screen "信号监控" 800x480, template "按钮"
   TextField "文本域_1" at 237,127 size 39x20; Text '状态'
   TextField "文本域_2" at 348,127 size 39x20; Text '地址'
   TextField "文本域_3" at 573,127 size 73x20; Text '注释名称'
   Group "Group" at 204,122 size 581x341
   TextField "文本域_30" at 240,127 size 39x20; Text '状态'
   Group "Group_1" at 204,122 size 581x341
   SymbolicIOField "符号 I/O 域_1" at 204,71 size 160x35; TextOn '1'; TextOff '0'; TextList "信号监控"
      on Change: ActivateScreenByNumber("跳转画面", 0)
      ProcessValue <- "跳转画面"
   GraphicView "图形视图_2" at 159,127 size 50x50; Picture "图形_2"
   Rectangle "矩形_2" at 207,152 size 109x15
      Appearance <- "操作面板急停"
   Rectangle "矩形_3" at 207,172 size 109x15
      Appearance <- "回原位"
   Rectangle "矩形_4" at 207,193 size 109x15
      Appearance <- "启动按钮"
   Rectangle "矩形_5" at 207,214 size 109x15
      Appearance <- "停止按钮"
   Rectangle "矩形_6" at 207,235 size 109x15
      Appearance <- "手动/自动"
   Rectangle "矩形_7" at 207,256 size 109x15
      Appearance <- "按钮盒急停"
   Rectangle "矩形_8" at 207,277 size 109x15
      Appearance <- "左启动"
   Rectangle "矩形_9" at 207,298 size 109x15
      Appearance <- "右启动"
   Rectangle "矩形_10" at 207,319 size 109x15
      Appearance <- "备用"
   Rectangle "矩形_11" at 207,340 size 109x15
      Appearance <- "安全光幕"
   Rectangle "矩形_12" at 207,361 size 109x15
      Appearance <- "Y1供料器有料"
   Rectangle "矩形_13" at 207,382 size 109x15
      Appearance <- "Y2供料器有料"
   Rectangle "矩形_14" at 207,403 size 109x15
      Appearance <- "1#工装产品信号"
   Rectangle "矩形_15" at 207,424 size 109x15
      Appearance <- "2#工装产品信号"
   TextField "文本域_4" at 348,150 size 41x20; Text 'I0.0'
   TextField "文本域_5" at 348,170 size 41x20; Text 'I0.1'
   TextField "文本域_6" at 348,191 size 41x20; Text 'I0.2'
   TextField "文本域_7" at 348,212 size 41x20; Text 'I0.3'
   TextField "文本域_8" at 348,233 size 41x20; Text 'I0.4'
   TextField "文本域_9" at 348,254 size 41x20; Text 'I0.5'
   TextField "文本域_10" at 348,275 size 41x20; Text 'I0.6'
   TextField "文本域_11" at 348,296 size 41x20; Text 'I0.7'
   TextField "文本域_12" at 348,317 size 41x20; Text 'I1.0'
   TextField "文本域_13" at 348,338 size 41x20; Text 'I1.1'
   TextField "文本域_14" at 348,359 size 41x20; Text 'I1.2'
   TextField "文本域_15" at 348,380 size 41x20; Text 'I1.3'
   TextField "文本域_16" at 348,401 size 41x20; Text 'I1.4'
   TextField "文本域_17" at 348,422 size 41x20; Text 'I1.5'
   TextField "文本域_18" at 561,151 size 101x19; Text '操作面板急停'
   TextField "文本域_19" at 561,171 size 85x19; Text '回原位按钮'
   TextField "文本域_20" at 561,192 size 101x19; Text '面板启动按钮'
   TextField "文本域_21" at 561,213 size 69x19; Text '停止按钮'
   TextField "文本域_22" at 561,234 size 78x19; Text '手动/自动'
   TextField "文本域_23" at 561,255 size 133x19; Text '双手启动面板急停'
   TextField "文本域_24" at 561,276 size 85x19; Text '左启动按钮'
   TextField "文本域_25" at 561,297 size 85x19; Text '右启动按钮'
   TextField "文本域_26" at 561,318 size 37x19; Text '备用'
   TextField "文本域_27" at 561,339 size 69x19; Text '光幕信号'
   TextField "文本域_28" at 561,360 size 103x19; Text 'Y1供料器有料'
   TextField "文本域_29" at 561,381 size 103x19; Text 'Y2供料器有料'
   TextField "文本域_31" at 561,402 size 119x19; Text '工装产品信号1#'
   TextField "文本域_32" at 561,423 size 119x19; Text '工装产品信号2#'

screen "I2.0" 800x480, template "按钮"
   Group "Group_1" at 204,122 size 581x341
   SymbolicIOField "符号 I/O 域_1" at 204,71 size 160x35; TextOn '1'; TextOff '0'; TextList "信号监控"
      on Change: ActivateScreenByNumber("跳转画面", 0)
      ProcessValue <- "跳转画面"
   GraphicView "图形视图_2" at 159,127 size 50x50; Picture "图形_2"
   Rectangle "矩形_2" at 207,152 size 109x15
      Appearance <- "气夹气缸到位2"
   Rectangle "矩形_3" at 207,172 size 109x15
      Appearance <- "气夹气缸到位1"
   Rectangle "矩形_4" at 207,193 size 109x15
      Appearance <- "工具错误"
   Rectangle "矩形_5" at 207,214 size 109x15
      Appearance <- "工具拧紧OK"
   Rectangle "矩形_6" at 207,235 size 109x15
      Appearance <- "工具拧紧NG"
   Rectangle "矩形_7" at 207,256 size 109x15
      Appearance <- "工具准备好"
   Rectangle "矩形_8" at 207,277 size 109x15
      Appearance <- "工具运行"
   Rectangle "矩形_9" at 207,298 size 109x15
      Appearance <- "气源压力检测"
   TextField "文本域_4" at 348,150 size 41x20; Text 'I2.0'
   TextField "文本域_5" at 348,170 size 41x20; Text 'I2.1'
   TextField "文本域_6" at 348,191 size 41x20; Text 'I2.2'
   TextField "文本域_7" at 348,212 size 41x20; Text 'I2.3'
   TextField "文本域_8" at 348,233 size 41x20; Text 'I2.4'
   TextField "文本域_9" at 348,254 size 41x20; Text 'I2.5'
   TextField "文本域_10" at 348,275 size 41x20; Text 'I2.6'
   TextField "文本域_11" at 348,296 size 41x20; Text 'I2.7'
   TextField "文本域_18" at 561,151 size 110x19; Text '气缸气夹到位2'
   TextField "文本域_19" at 561,171 size 110x19; Text '气缸气夹到位1'
   TextField "文本域_20" at 561,192 size 69x19; Text '工具错误'
   TextField "文本域_21" at 561,213 size 87x19; Text '工具拧紧OK'
   TextField "文本域_22" at 561,234 size 87x19; Text '工具拧紧NG'
   TextField "文本域_23" at 561,255 size 85x19; Text '工具准备好'
   TextField "文本域_24" at 561,276 size 69x19; Text '工具运行'
   TextField "文本域_25" at 561,297 size 101x19; Text '气源压力检测'
   Group "Group" at 204,122 size 581x341
   TextField "文本域_30" at 240,127 size 39x20; Text '状态'
   TextField "文本域_1" at 237,127 size 39x20; Text '状态'
   TextField "文本域_2" at 348,127 size 39x20; Text '地址'
   TextField "文本域_3" at 573,127 size 73x20; Text '注释名称'

screen "I3.0" 800x480, template "按钮"
   Group "Group_1" at 204,122 size 581x341
   SymbolicIOField "符号 I/O 域_1" at 204,71 size 160x35; TextOn '1'; TextOff '0'; TextList "信号监控"
      on Change: ActivateScreenByNumber("跳转画面", 0)
      ProcessValue <- "跳转画面"
   GraphicView "图形视图_2" at 159,127 size 50x50; Picture "图形_2"
   Rectangle "矩形_2" at 207,152 size 109x15
      Appearance <- "光栅屏蔽对射开关"
   Rectangle "矩形_3" at 207,172 size 109x15
      Appearance <- "吸附信号"
   Rectangle "矩形_4" at 207,193 size 109x15
      Appearance <- "电批下压气缸信号"
   Rectangle "矩形_5" at 207,214 size 109x15
      Appearance <- "安全门"
   Rectangle "矩形_6" at 207,235 size 109x15
      Appearance <- "回原位中"
   Rectangle "矩形_7" at 207,256 size 109x15
      Appearance <- "回原位完成"
   Rectangle "矩形_8" at 207,277 size 109x15
      Appearance <- "X轴故障报警"
   Rectangle "矩形_9" at 207,298 size 109x15
      Appearance <- "Y轴故障报警"
   TextField "文本域_4" at 348,150 size 41x20; Text 'I3.0'
   TextField "文本域_5" at 348,170 size 41x20; Text 'I3.1'
   TextField "文本域_6" at 348,191 size 41x20; Text 'I3.2'
   TextField "文本域_7" at 348,212 size 41x20; Text 'I3.3'
   TextField "文本域_8" at 348,233 size 41x20; Text 'I3.4'
   TextField "文本域_9" at 348,254 size 41x20; Text 'I3.5'
   TextField "文本域_10" at 348,275 size 41x20; Text 'I3.6'
   TextField "文本域_11" at 348,296 size 41x20; Text 'I3.7'
   TextField "文本域_18" at 561,151 size 101x19; Text '光栅屏蔽开关'
   TextField "文本域_19" at 561,171 size 69x19; Text '吸附信号'
   TextField "文本域_20" at 561,192 size 133x19; Text '电批下压气缸信号'
   TextField "文本域_21" at 561,213 size 53x19; Text '安全门'
   TextField "文本域_22" at 561,234 size 53x19; Text '回原位'
   TextField "文本域_23" at 561,255 size 85x19; Text '回原位完成'
   TextField "文本域_24" at 561,276 size 94x19; Text 'X轴伺服报警'
   TextField "文本域_25" at 561,297 size 94x19; Text 'Y轴伺服报警'
   Group "Group" at 204,122 size 581x341
   TextField "文本域_30" at 240,127 size 39x20; Text '状态'
   TextField "文本域_1" at 237,127 size 39x20; Text '状态'
   TextField "文本域_2" at 348,127 size 39x20; Text '地址'
   TextField "文本域_3" at 573,127 size 73x20; Text '注释名称'

screen "I4.0" 800x480, template "按钮"
   Group "Group_1" at 204,122 size 581x341
   SymbolicIOField "符号 I/O 域_1" at 204,71 size 160x35; TextOn '1'; TextOff '0'; TextList "信号监控"
      on Change: ActivateScreenByNumber("跳转画面", 0)
      ProcessValue <- "跳转画面"
   GraphicView "图形视图_2" at 159,127 size 50x50; Picture "图形_2"
   Rectangle "矩形_2" at 207,152 size 109x15
      Appearance <- "Z轴故障报警"
   Rectangle "矩形_3" at 207,172 size 109x15
      Appearance <- "运动控制卡完成/释放夹紧气缸"
   Rectangle "矩形_4" at 207,193 size 109x15
      Appearance <- "备用_3"
   Rectangle "矩形_5" at 207,214 size 109x15
      Appearance <- "备用_4"
   Rectangle "矩形_6" at 207,235 size 109x15
      Appearance <- "备用_5"
   Rectangle "矩形_7" at 207,256 size 109x15
      Appearance <- "备用_6"
   Rectangle "矩形_8" at 207,277 size 109x15
      Appearance <- "备用_7"
   Rectangle "矩形_9" at 207,298 size 109x15
      Appearance <- "备用_8"
   TextField "文本域_4" at 348,150 size 41x20; Text 'I4.0'
   TextField "文本域_5" at 348,170 size 41x20; Text 'I4.1'
   TextField "文本域_6" at 348,191 size 41x20; Text 'I4.2'
   TextField "文本域_7" at 348,212 size 41x20; Text 'I4.3'
   TextField "文本域_8" at 348,233 size 41x20; Text 'I4.4'
   TextField "文本域_9" at 348,254 size 41x20; Text 'I4.5'
   TextField "文本域_10" at 348,275 size 41x20; Text 'I4.6'
   TextField "文本域_11" at 348,296 size 41x20; Text 'I4.7'
   TextField "文本域_18" at 561,151 size 94x19; Text 'Z轴伺服报警'
   TextField "文本域_19" at 561,171 size 133x19; Text '运动控制完成信号'
   TextField "文本域_20" at 561,192 size 37x19; Text '备用'
   TextField "文本域_21" at 561,213 size 37x19; Text '备用'
   TextField "文本域_22" at 561,234 size 37x19; Text '备用'
   TextField "文本域_23" at 561,255 size 37x19; Text '备用'
   TextField "文本域_24" at 561,276 size 37x19; Text '备用'
   TextField "文本域_25" at 561,297 size 37x19; Text '备用'
   Group "Group" at 204,122 size 581x341
   TextField "文本域_30" at 240,127 size 39x20; Text '状态'
   TextField "文本域_1" at 237,127 size 39x20; Text '状态'
   TextField "文本域_2" at 348,127 size 39x20; Text '地址'
   TextField "文本域_3" at 573,127 size 73x20; Text '注释名称'

screen "Q0.0" 800x480, template "按钮"
   Group "Group_1" at 204,122 size 581x341
   SymbolicIOField "符号 I/O 域_1" at 204,71 size 160x35; TextOn '1'; TextOff '0'; TextList "信号监控"
      on Change: ActivateScreenByNumber("跳转画面", 0)
      ProcessValue <- "跳转画面"
   GraphicView "图形视图_2" at 159,127 size 50x50; Picture "图形_2"
   Rectangle "矩形_2" at 207,152 size 109x15
      Appearance <- "三色灯黄色"
   Rectangle "矩形_3" at 207,172 size 109x15
      Appearance <- "三色灯绿色"
   Rectangle "矩形_4" at 207,193 size 109x15
      Appearance <- "三色灯红色"
   Rectangle "矩形_5" at 207,214 size 109x15
      Appearance <- "三色灯蜂鸣器"
   Rectangle "矩形_6" at 207,235 size 109x15
      Appearance <- "绿色半球指示灯"
   Rectangle "矩形_7" at 207,256 size 109x15
      Appearance <- "红色半球指示灯"
   Rectangle "矩形_8" at 207,277 size 109x15
      Appearance <- "运动控制卡任务选择1"
   Rectangle "矩形_9" at 207,298 size 109x15
      Appearance <- "运动控制卡任务选择2"
   Rectangle "矩形_10" at 207,319 size 109x15
      Appearance <- "运动控制卡任务选择3"
   Rectangle "矩形_11" at 207,340 size 109x15
      Appearance <- "运动控制卡任务选择4"
   TextField "文本域_4" at 348,150 size 41x20; Text 'Q0.0'
   TextField "文本域_5" at 348,170 size 41x20; Text 'Q0.1'
   TextField "文本域_6" at 348,191 size 41x20; Text 'Q0.2'
   TextField "文本域_7" at 348,212 size 41x20; Text 'Q0.3'
   TextField "文本域_8" at 348,233 size 41x20; Text 'Q0.4'
   TextField "文本域_9" at 348,254 size 41x20; Text 'Q0.5'
   TextField "文本域_10" at 348,275 size 41x20; Text 'Q0.6'
   TextField "文本域_11" at 348,296 size 41x20; Text 'Q0.7'
   TextField "文本域_12" at 348,317 size 41x20; Text 'Q1.0'
   TextField "文本域_13" at 348,338 size 41x20; Text 'Q1.1'
   TextField "文本域_18" at 561,151 size 69x19; Text '三色灯黄'
   TextField "文本域_19" at 561,171 size 69x19; Text '三色灯绿'
   TextField "文本域_20" at 561,192 size 69x19; Text '三色灯红'
   TextField "文本域_21" at 561,213 size 101x19; Text '三色灯蜂鸣器'
   TextField "文本域_22" at 561,234 size 101x19; Text '半球指示灯绿'
   TextField "文本域_23" at 561,255 size 101x19; Text '半球指示灯红'
   TextField "文本域_24" at 561,276 size 174x19; Text '运动控制板卡任务选择1'
   TextField "文本域_25" at 561,297 size 174x19; Text '运动控制板卡任务选择2'
   TextField "文本域_26" at 561,318 size 174x19; Text '运动控制板卡任务选择3'
   TextField "文本域_27" at 561,339 size 174x19; Text '运动控制板卡任务选择4'
   Group "Group" at 204,122 size 581x341
   TextField "文本域_30" at 240,127 size 39x20; Text '状态'
   TextField "文本域_1" at 237,127 size 39x20; Text '状态'
   TextField "文本域_2" at 348,127 size 39x20; Text '地址'
   TextField "文本域_3" at 573,127 size 73x20; Text '注释名称'

screen "Q2.0" 800x480, template "按钮"
   Group "Group_1" at 204,122 size 581x341
   SymbolicIOField "符号 I/O 域_1" at 204,71 size 160x35; TextOn '1'; TextOff '0'; TextList "信号监控"
      on Change: ActivateScreenByNumber("跳转画面", 0)
      ProcessValue <- "跳转画面"
   GraphicView "图形视图_2" at 159,127 size 50x50; Picture "图形_2"
   Rectangle "矩形_2" at 207,152 size 109x15
      Appearance <- "运动控制卡任务选择5"
   Rectangle "矩形_3" at 207,172 size 109x15
      Appearance <- "Y1供料器有料输出"
   Rectangle "矩形_4" at 207,193 size 109x15
      Appearance <- "Y2供料器有料输出"
   Rectangle "矩形_5" at 207,214 size 109x15
      Appearance <- "运动控制卡启动"
   Rectangle "矩形_6" at 207,235 size 109x15
      Appearance <- "运动控制卡复位"
   Rectangle "矩形_7" at 207,256 size 109x15
      Appearance <- "电批急停"
   Rectangle "矩形_8" at 207,277 size 109x15
      Appearance <- "运动控制卡停止"
   Rectangle "矩形_9" at 207,298 size 109x15
      Appearance <- "吸取螺丝电磁阀"
   TextField "文本域_4" at 348,150 size 41x20; Text 'Q2.0'
   TextField "文本域_5" at 348,170 size 41x20; Text 'Q2.1'
   TextField "文本域_6" at 348,191 size 41x20; Text 'Q2.2'
   TextField "文本域_7" at 348,212 size 41x20; Text 'Q2.3'
   TextField "文本域_8" at 348,233 size 41x20; Text 'Q2.4'
   TextField "文本域_9" at 348,254 size 41x20; Text 'Q2.5'
   TextField "文本域_10" at 348,275 size 41x20; Text 'Q2.6'
   TextField "文本域_11" at 348,296 size 41x20; Text 'Q2.7'
   TextField "文本域_18" at 561,151 size 174x19; Text '运动控制板卡任务选择5'
   TextField "文本域_19" at 561,171 size 103x19; Text 'Y1供料器有料'
   TextField "文本域_20" at 561,192 size 103x19; Text 'Y2供料器有料'
   TextField "文本域_21" at 561,213 size 69x19; Text '设备启动'
   TextField "文本域_22" at 561,234 size 53x19; Text '回原位'
   TextField "文本域_23" at 561,255 size 69x19; Text '紧急停止'
   TextField "文本域_24" at 561,276 size 69x19; Text '设备停止'
   TextField "文本域_25" at 561,297 size 117x19; Text '吸取螺丝电磁阀'
   Group "Group" at 204,122 size 581x341
   TextField "文本域_30" at 240,127 size 39x20; Text '状态'
   TextField "文本域_1" at 237,127 size 39x20; Text '状态'
   TextField "文本域_2" at 348,127 size 39x20; Text '地址'
   TextField "文本域_3" at 573,127 size 73x20; Text '注释名称'

screen "Q3.0" 800x480, template "按钮"
   Group "Group_1" at 204,122 size 581x341
   SymbolicIOField "符号 I/O 域_1" at 204,71 size 160x35; TextOn '1'; TextOff '0'; TextList "信号监控"
      on Change: ActivateScreenByNumber("跳转画面", 0)
      ProcessValue <- "跳转画面"
   GraphicView "图形视图_2" at 159,127 size 50x50; Picture "图形_2"
   Rectangle "矩形_2" at 207,152 size 109x15
      Appearance <- "下压气缸电磁阀"
   Rectangle "矩形_3" at 207,172 size 109x15
      Appearance <- "工装电磁铁"
   Rectangle "矩形_4" at 207,193 size 109x15
      Appearance <- "运动控制光栅报警"
   Rectangle "矩形_5" at 207,214 size 109x15
      Appearance <- "伺服复位"
   Rectangle "矩形_6" at 207,235 size 109x15
      Appearance <- "电批急停"
   Rectangle "矩形_7" at 207,256 size 109x15
      Appearance <- "备用_3(1)"
   Rectangle "矩形_8" at 207,277 size 109x15
      Appearance <- "FFU"
   Rectangle "矩形_9" at 207,298 size 109x15
      Appearance <- "照明"
   TextField "文本域_4" at 348,150 size 41x20; Text 'Q3.0'
   TextField "文本域_5" at 348,170 size 41x20; Text 'Q3.1'
   TextField "文本域_6" at 348,191 size 41x20; Text 'Q3.2'
   TextField "文本域_7" at 348,212 size 41x20; Text 'Q3.3'
   TextField "文本域_8" at 348,233 size 41x20; Text 'Q3.4'
   TextField "文本域_9" at 348,254 size 41x20; Text 'Q3.5'
   TextField "文本域_10" at 348,275 size 41x20; Text 'Q3.6'
   TextField "文本域_11" at 348,296 size 41x20; Text 'Q3.7'
   TextField "文本域_18" at 561,151 size 117x19; Text '下压气缸电磁阀'
   TextField "文本域_19" at 561,171 size 53x19; Text '电磁铁'
   TextField "文本域_20" at 561,192 size 69x19; Text '光幕报警'
   TextField "文本域_21" at 561,213 size 69x19; Text '伺服复位'
   TextField "文本域_22" at 561,234 size 69x19; Text '电批急停'
   TextField "文本域_23" at 561,255 size 101x19; Text '电批测试启动'
   TextField "文本域_24" at 562,276 size 32x19; Text 'FFU'
   TextField "文本域_25" at 561,297 size 37x19; Text '照明'
   Group "Group" at 204,122 size 581x341
   TextField "文本域_30" at 240,127 size 39x20; Text '状态'
   TextField "文本域_1" at 237,127 size 39x20; Text '状态'
   TextField "文本域_2" at 348,127 size 39x20; Text '地址'
   TextField "文本域_3" at 573,127 size 73x20; Text '注释名称'

screen "Q4.0" 800x480, template "按钮"
   Group "Group_1" at 204,122 size 581x341
   SymbolicIOField "符号 I/O 域_1" at 204,71 size 160x35; TextOn '1'; TextOff '0'; TextList "信号监控"
      on Change: ActivateScreenByNumber("跳转画面", 0)
      ProcessValue <- "跳转画面"
   GraphicView "图形视图_2" at 159,127 size 50x50; Picture "图形_2"
   Rectangle "矩形_2" at 207,152 size 109x15
      Appearance <- "夹紧气缸1夹紧"
   Rectangle "矩形_3" at 207,172 size 109x15
      Appearance <- "夹紧气缸2夹紧"
   Rectangle "矩形_4" at 207,193 size 109x15
      Appearance <- "备用_3(1)"
   Rectangle "矩形_5" at 207,214 size 109x15
      Appearance <- "备用_4(1)"
   Rectangle "矩形_6" at 207,235 size 109x15
      Appearance <- "备用_5(1)"
   Rectangle "矩形_7" at 207,256 size 109x15
      Appearance <- "备用_6(1)"
   Rectangle "矩形_8" at 207,277 size 109x15
      Appearance <- "备用_7(1)"
   Rectangle "矩形_9" at 207,298 size 109x15
      Appearance <- "备用_8(1)"
   TextField "文本域_4" at 348,150 size 41x20; Text 'Q4.0'
   TextField "文本域_5" at 348,170 size 41x20; Text 'Q4.1'
   TextField "文本域_6" at 348,191 size 41x20; Text 'Q4.2'
   TextField "文本域_7" at 348,212 size 41x20; Text 'Q4.3'
   TextField "文本域_8" at 348,233 size 41x20; Text 'Q4.4'
   TextField "文本域_9" at 348,254 size 41x20; Text 'Q4.5'
   TextField "文本域_10" at 348,275 size 41x20; Text 'Q4.6'
   TextField "文本域_11" at 348,296 size 41x20; Text 'Q4.7'
   TextField "文本域_18" at 561,151 size 101x19; Text '左启动按钮灯'
   TextField "文本域_19" at 561,171 size 101x19; Text '右启动按钮灯'
   TextField "文本域_20" at 561,192 size 69x19; Text '气缸夹紧'
   TextField "文本域_21" at 561,213 size 37x19; Text '备用'
   TextField "文本域_22" at 561,234 size 37x19; Text '备用'
   TextField "文本域_23" at 561,255 size 37x19; Text '备用'
   TextField "文本域_24" at 561,276 size 37x19; Text '备用'
   TextField "文本域_25" at 561,297 size 37x19; Text '备用'
   Group "Group" at 204,122 size 581x341
   TextField "文本域_30" at 240,127 size 39x20; Text '状态'
   TextField "文本域_1" at 237,127 size 39x20; Text '状态'
   TextField "文本域_2" at 348,127 size 39x20; Text '地址'
   TextField "文本域_3" at 573,127 size 73x20; Text '注释名称'

screen "X1" 800x480, template "按钮"
   Group "Group_1" at 204,122 size 581x341
   SymbolicIOField "符号 I/O 域_1" at 204,71 size 160x35; TextOn '1'; TextOff '0'; TextList "信号监控"
      on Change: ActivateScreenByNumber("跳转画面", 0)
      ProcessValue <- "跳转画面"
   GraphicView "图形视图_2" at 159,127 size 50x50; Picture "图形_2"
   Rectangle "矩形_2" at 207,152 size 109x15
      Appearance <- "HengKongMC_输入_X轴原位"
   Rectangle "矩形_3" at 207,172 size 109x15
      Appearance <- "HengKongMC_输入_Y轴原位"
   Rectangle "矩形_4" at 207,193 size 109x15
      Appearance <- "HengKongMC_输入_Z轴原位"
   Rectangle "矩形_5" at 207,214 size 109x15
      Appearance <- "HengKongMC_输入_X4备用"
   Rectangle "矩形_6" at 207,235 size 109x15
      Appearance <- "HengKongMC_输入_Y2供料器有料"
   Rectangle "矩形_7" at 207,256 size 109x15
      Appearance <- "HengKongMC_输入_电批启动"
   Rectangle "矩形_8" at 207,277 size 109x15
      Appearance <- "HengKongMC_输入_任务选择1"
   Rectangle "矩形_9" at 207,298 size 109x15
      Appearance <- "HengKongMC_输入_任务选择2"
   TextField "文本域_4" at 348,150 size 23x20; Text 'X1'
   TextField "文本域_5" at 348,170 size 23x20; Text 'X2'
   TextField "文本域_6" at 348,191 size 23x20; Text 'X3'
   TextField "文本域_7" at 348,212 size 23x20; Text 'X4'
   TextField "文本域_8" at 348,233 size 23x20; Text 'X5'
   TextField "文本域_9" at 348,254 size 23x20; Text 'X6'
   TextField "文本域_10" at 348,275 size 23x20; Text 'X7'
   TextField "文本域_11" at 348,296 size 23x20; Text 'X8'
   TextField "文本域_18" at 561,151 size 94x19; Text 'X轴原位信号'
   TextField "文本域_19" at 561,171 size 94x19; Text 'Y轴原位信号'
   TextField "文本域_20" at 561,192 size 94x19; Text 'Z轴原位信号'
   TextField "文本域_21" at 561,213 size 37x19; Text '备用'
   TextField "文本域_22" at 561,234 size 103x19; Text 'Y2供料器有料'
   TextField "文本域_23" at 561,255 size 69x19; Text '电批启动'
   TextField "文本域_24" at 561,276 size 78x19; Text '任务选择1'
   TextField "文本域_25" at 561,297 size 78x19; Text '任务选择2'
   TextField "文本域_12" at 348,317 size 23x20; Text 'X9'
   TextField "文本域_13" at 348,338 size 32x20; Text 'X10'
   TextField "文本域_14" at 348,359 size 32x20; Text 'X11'
   TextField "文本域_15" at 348,380 size 32x20; Text 'X12'
   TextField "文本域_16" at 348,401 size 32x20; Text 'X13'
   TextField "文本域_17" at 348,422 size 32x20; Text 'X14'
   TextField "文本域_26" at 348,443 size 32x20; Text 'X15'
   TextField "文本域_27" at 561,318 size 37x19; Text '启动'
   TextField "文本域_28" at 561,339 size 53x19; Text '回原位'
   TextField "文本域_29" at 561,360 size 37x19; Text '急停'
   TextField "文本域_31" at 561,381 size 55x19; Text '电批OK'
   TextField "文本域_32" at 561,402 size 69x19; Text '光栅报警'
   TextField "文本域_33" at 561,423 size 78x19; Text '任务选择3'
   TextField "文本域_34" at 561,444 size 78x19; Text '任务选择4'
   Rectangle "矩形_10" at 207,318 size 109x15
      Appearance <- "HengKongMC_输入_启动"
   Rectangle "矩形_11" at 207,339 size 109x15
      Appearance <- "HengKongMC_输入_回原位"
   Rectangle "矩形_12" at 207,360 size 109x15
      Appearance <- "HengKongMC_输入_急停"
   Rectangle "矩形_13" at 207,381 size 109x15
      Appearance <- "HengKongMC_输入_OK"
   Rectangle "矩形_14" at 207,402 size 109x15
      Appearance <- "HengKongMC_输入_光幕和门控报警"
   Rectangle "矩形_15" at 207,423 size 109x15
      Appearance <- "HengKongMC_输入_任务选择3"
   Rectangle "矩形_16" at 207,444 size 109x15
      Appearance <- "HengKongMC_输入_任务选择4"
   Group "Group" at 204,122 size 581x341
   TextField "文本域_30" at 240,127 size 39x20; Text '状态'
   TextField "文本域_1" at 237,127 size 39x20; Text '状态'
   TextField "文本域_2" at 348,127 size 39x20; Text '地址'
   TextField "文本域_3" at 573,127 size 73x20; Text '注释名称'

screen "X16" 800x480, template "按钮"
   Group "Group_1" at 204,122 size 581x341
   SymbolicIOField "符号 I/O 域_1" at 204,71 size 160x35; TextOn '1'; TextOff '0'; TextList "信号监控"
      on Change: ActivateScreenByNumber("跳转画面", 0)
      ProcessValue <- "跳转画面"
   GraphicView "图形视图_2" at 159,127 size 50x50; Picture "图形_2"
   Rectangle "矩形_2" at 207,152 size 109x15
      Appearance <- "HengKongMC_输入_任务选择5"
   Rectangle "矩形_3" at 207,172 size 109x15
      Appearance <- "HengKongMC_输入_负压传感器"
   Rectangle "矩形_4" at 207,193 size 109x15
      Appearance <- "HengKongMC_输入_Y1供料器有料"
   Rectangle "矩形_5" at 207,214 size 109x15
      Appearance <- "HengKongMC_输入_X19"
   Rectangle "矩形_6" at 207,235 size 109x15
      Appearance <- "HengKongMC_输入_X20"
   Rectangle "矩形_7" at 207,256 size 109x15
      Appearance <- "HengKongMC_输入_X21"
   Rectangle "矩形_8" at 207,277 size 109x15
      Appearance <- "HengKongMC_输入_下压气缸原位"
   Rectangle "矩形_9" at 207,298 size 109x15
      Appearance <- "HengKongMC_输入_X23"
   TextField "文本域_4" at 348,150 size 32x20; Text 'X16'
   TextField "文本域_5" at 348,170 size 32x20; Text 'X17'
   TextField "文本域_6" at 348,191 size 32x20; Text 'X18'
   TextField "文本域_7" at 348,212 size 32x20; Text 'X19'
   TextField "文本域_8" at 348,233 size 32x20; Text 'X20'
   TextField "文本域_9" at 348,254 size 32x20; Text 'X21'
   TextField "文本域_10" at 348,275 size 32x20; Text 'X22'
   TextField "文本域_11" at 348,296 size 32x20; Text 'X23'
   TextField "文本域_18" at 561,151 size 78x19; Text '任务选择5'
   TextField "文本域_19" at 561,171 size 85x19; Text '负压传感器'
   TextField "文本域_20" at 561,192 size 103x19; Text 'Y1供料器有料'
   TextField "文本域_21" at 561,213 size 37x19; Text '备用'
   TextField "文本域_22" at 561,234 size 37x19; Text '备用'
   TextField "文本域_23" at 561,255 size 37x19; Text '备用'
   TextField "文本域_24" at 561,276 size 101x19; Text '下压气缸原位'
   TextField "文本域_25" at 561,297 size 37x19; Text '备用'
   TextField "文本域_12" at 348,317 size 32x20; Text 'X24'
   TextField "文本域_27" at 561,318 size 37x19; Text '停止'
   Rectangle "矩形_10" at 207,318 size 109x15
      Appearance <- "HengKongMC_输入_停止"
   Group "Group" at 204,122 size 581x341
   TextField "文本域_30" at 240,127 size 39x20; Text '状态'
   TextField "文本域_1" at 237,127 size 39x20; Text '状态'
   TextField "文本域_2" at 348,127 size 39x20; Text '地址'
   TextField "文本域_3" at 573,127 size 73x20; Text '注释名称'

screen "Y1" 800x480, template "按钮"
   Group "Group_1" at 204,122 size 581x341
   SymbolicIOField "符号 I/O 域_1" at 204,71 size 160x35; TextOn '1'; TextOff '0'; TextList "信号监控"
      on Change: ActivateScreenByNumber("跳转画面", 0)
      ProcessValue <- "跳转画面"
   GraphicView "图形视图_2" at 159,127 size 50x50; Picture "图形_2"
   Rectangle "矩形_2" at 207,152 size 109x15
      Appearance <- "HengKongMC_输出_吸取螺丝信号"
   Rectangle "矩形_3" at 207,172 size 109x15
      Appearance <- "HengKongMC_输出_回原位成功"
   Rectangle "矩形_4" at 207,193 size 109x15
      Appearance <- "HengKongMC_输出_回原位中"
   Rectangle "矩形_5" at 207,214 size 109x15
      Appearance <- "HengKongMC_输出_下压气缸信号"
   Rectangle "矩形_6" at 207,235 size 109x15
      Appearance <- "HengKongMC_输出_Y5"
   Rectangle "矩形_7" at 207,256 size 109x15
      Appearance <- "HengKongMC_输出_认螺帽反转"
   Rectangle "矩形_8" at 207,277 size 109x15
      Appearance <- "HengKongMC_输出_Y7"
   Rectangle "矩形_9" at 207,298 size 109x15
      Appearance <- "HengKongMC_输出_Y8"
   TextField "文本域_4" at 348,150 size 23x20; Text 'Y1'
   TextField "文本域_5" at 348,170 size 23x20; Text 'Y2'
   TextField "文本域_6" at 348,191 size 23x20; Text 'Y3'
   TextField "文本域_7" at 348,212 size 23x20; Text 'Y4'
   TextField "文本域_8" at 348,233 size 23x20; Text 'Y5'
   TextField "文本域_9" at 348,254 size 23x20; Text 'Y6'
   TextField "文本域_10" at 348,275 size 23x20; Text 'Y7'
   TextField "文本域_11" at 348,296 size 23x20; Text 'Y8'
   TextField "文本域_18" at 561,151 size 101x19; Text '吸取螺丝信号'
   TextField "文本域_19" at 561,171 size 85x19; Text '回原位成功'
   TextField "文本域_20" at 561,192 size 69x19; Text '回原位中'
   TextField "文本域_21" at 561,213 size 133x19; Text '下压气缸下压信号'
   TextField "文本域_22" at 561,234 size 37x19; Text '备用'
   TextField "文本域_23" at 561,255 size 85x19; Text '认螺帽反转'
   TextField "文本域_24" at 561,276 size 149x19; Text '运动控制卡完成信号'
   TextField "文本域_25" at 561,297 size 37x19; Text '备用'
   TextField "文本域_12" at 348,317 size 23x20; Text 'Y9'
   TextField "文本域_13" at 348,338 size 32x20; Text 'Y10'
   TextField "文本域_14" at 348,359 size 32x20; Text 'Y11'
   TextField "文本域_15" at 348,380 size 32x20; Text 'Y12'
   TextField "文本域_16" at 348,401 size 32x20; Text 'Y13'
   TextField "文本域_17" at 348,422 size 32x20; Text 'Y14'
   TextField "文本域_26" at 348,443 size 32x20; Text 'Y15'
   TextField "文本域_27" at 561,318 size 78x19; Text '电批任务0'
   TextField "文本域_28" at 561,339 size 78x19; Text '电批任务1'
   TextField "文本域_29" at 561,360 size 78x19; Text '电批任务2'
   TextField "文本域_31" at 561,381 size 37x19; Text '备用'
   TextField "文本域_32" at 561,402 size 69x19; Text '启动电批'
   TextField "文本域_33" at 561,423 size 37x19; Text '备用'
   TextField "文本域_34" at 561,444 size 101x19; Text '回原位标志位'
   Rectangle "矩形_10" at 207,318 size 109x15
      Appearance <- "HengKongMC_输出_任务选择0"
   Rectangle "矩形_11" at 207,339 size 109x15
      Appearance <- "HengKongMC_输出_任务选择1"
   Rectangle "矩形_12" at 207,360 size 109x15
      Appearance <- "HengKongMC_输出_任务选择2"
   Rectangle "矩形_13" at 207,381 size 109x15
      Appearance <- "HengKongMC_输出_Y12"
   Rectangle "矩形_14" at 207,402 size 109x15
      Appearance <- "HengKongMC_输出_启动电批"
   Rectangle "矩形_15" at 207,423 size 109x15
      Appearance <- "HengKongMC_输出_Y14"
   Rectangle "矩形_16" at 207,444 size 109x15
      Appearance <- "回原位标志位"
   Group "Group" at 204,122 size 581x341
   TextField "文本域_30" at 240,127 size 39x20; Text '状态'
   TextField "文本域_1" at 237,127 size 39x20; Text '状态'
   TextField "文本域_2" at 348,127 size 39x20; Text '地址'
   TextField "文本域_3" at 573,127 size 73x20; Text '注释名称'

screen "Y16" 800x480, template "按钮"
   Group "Group_1" at 204,122 size 581x341
   SymbolicIOField "符号 I/O 域_1" at 204,71 size 160x35; TextOn '1'; TextOff '0'; TextList "信号监控"
      on Change: ActivateScreenByNumber("跳转画面", 0)
      ProcessValue <- "跳转画面"
   GraphicView "图形视图_2" at 159,127 size 50x50; Picture "图形_2"
   Rectangle "矩形_2" at 207,152 size 109x15
      Appearance <- "HengKongMC_输出_Y16"
   TextField "文本域_4" at 348,150 size 32x20; Text 'Y16'
   TextField "文本域_18" at 561,151 size 37x19; Text '备用'
   Group "Group" at 204,122 size 581x341
   TextField "文本域_30" at 240,127 size 39x20; Text '状态'
   TextField "文本域_1" at 237,127 size 39x20; Text '状态'
   TextField "文本域_2" at 348,127 size 39x20; Text '地址'
   TextField "文本域_3" at 573,127 size 73x20; Text '注释名称'

screen "屏蔽管理" 800x480, template "按钮"
   TextField "文本域_3" at 639,76 size 73x20; Text '操作按钮'
   TextField "文本域_2" at 421,76 size 73x20; Text '注释名称'
   Group "Group" at 359,67 size 422x401
   GraphicView "图形视图_2" at 159,305 size 50x50; Picture "图形_2"
   TextField "文本域_6" at 375,122 size 167x23; Text 'Y1供料器报警屏蔽'
   TextField "文本域_4" at 375,174 size 167x23; Text 'Y2供料器报警屏蔽'
   TextField "文本域_5" at 375,226 size 176x23; Text '工装产品检测1屏蔽'
   TextField "文本域_7" at 375,278 size 176x23; Text '工装产品检测2屏蔽'
   TextField "文本域_8" at 410,381 size 16x23; Text 'Text'
   TextField "文本域_10" at 375,330 size 165x23; Text '工装夹紧气缸屏蔽'
   SymbolicIOField "符号 I/O 域_1" at 595,113 size 157x32; TextOff '0'; TextOn '1'; TextList "屏蔽信号"
      ProcessValue <- "Blocking function_Y1供料器报警屏蔽"
   TextField "文本域_11" at 375,434 size 185x23; Text '上位机启动信号屏蔽'
   SymbolicIOField "符号 I/O 域_2" at 595,165 size 157x32; TextOn '1'; TextOff '0'; TextList "屏蔽信号"
      ProcessValue <- "Blocking function_Y2供料器报警屏蔽"
   SymbolicIOField "符号 I/O 域_3" at 595,218 size 157x32; TextOn '1'; TextOff '0'; TextList "屏蔽信号"
      ProcessValue <- "Blocking function_工装产品检测1屏蔽"
   SymbolicIOField "符号 I/O 域_4" at 595,271 size 157x32; TextOn '1'; TextOff '0'; TextList "屏蔽信号"
      ProcessValue <- "Blocking function_工装产品检测2屏蔽"
   SymbolicIOField "符号 I/O 域_5" at 595,324 size 157x32; TextOn '1'; TextOff '0'; TextList "屏蔽信号"
      ProcessValue <- "Blocking function_夹紧气缸1夹紧屏蔽"
   SymbolicIOField "符号 I/O 域_6" at 595,377 size 157x32; TextOn '1'; TextOff '0'; TextList "屏蔽信号"
      ProcessValue <- "Blocking function_夹紧气缸2夹紧屏蔽"
   SymbolicIOField "符号 I/O 域_7" at 595,430 size 157x32; TextOn '1'; TextOff '0'; TextList "屏蔽信号"
      ProcessValue <- "Blocking function_上位机屏蔽"
   TextField "文本域_9" at 375,382 size 165x23; Text '工装夹紧气缸屏蔽'
   SymbolicIOField "符号 I/O 域_8" at 185,69 size 160x35; TextOn '1'; TextOff '0'; TextList "屏蔽菜单"
      ProcessValue <- "屏蔽菜单"
      on Change: ActivateScreenByNumber("屏蔽菜单", 0)

screen "伺服状态" 800x480, template "按钮"
   GraphicView "图形视图_1" at 295,87 size 51x51; Picture "图形_19"
      Visibility <- "准备OKx"
   GraphicView "图形视图_2" at 295,87 size 51x51; Picture "图形_20"
      Visibility <- "准备OKx"
   GraphicView "图形视图_3" at 295,293 size 51x51; Picture "图形_19"
      Visibility <- "准备OKy"
   GraphicView "图形视图_4" at 295,293 size 51x51; Picture "图形_20"
      Visibility <- "准备OKy"
   GraphicView "图形视图_5" at 625,162 size 51x51; Picture "图形_19"
      Visibility <- "准备OKz"
   GraphicView "图形视图_6" at 625,162 size 51x51; Picture "图形_20"
      Visibility <- "准备OKz"
   Rectangle "矩形_1" at 280,158 size 14x40
      Appearance <- "正方向x"
   Rectangle "矩形_2" at 225,222 size 14x40
      Appearance <- "正方向y"
   Rectangle "矩形_3" at 548,82 size 14x40
      Appearance <- "正方向z"
   Rectangle "矩形_4" at 718,158 size 14x40
      Appearance <- "负方向x"
   Rectangle "矩形_5" at 225,400 size 14x40
      Appearance <- "负方向y"
   Rectangle "矩形_6" at 548,272 size 14x40
      Appearance <- "负方向z"
   GraphicView "图形视图_7" at 159,367 size 50x50; Picture "图形_2"
   TextField "文本域_1" at 214,84 size 45x29; Text 'X轴'
   TextField "文本域_2" at 296,227 size 45x29; Text 'Y轴'
   TextField "文本域_3" at 646,93 size 45x29; Text 'Z轴'
   TextField "文本域_4" at 601,375 size 19x29; Text 'Text'
   TextField "文本域_5" at 562,356 size 73x20; Text '限位正常'
   GraphicView "图形视图_8" at 640,404 size 51x51; Picture "图形_20"
   TextField "文本域_6" at 703,420 size 73x20; Text '故障报警'
   GraphicView "图形视图_9" at 505,404 size 51x51; Picture "图形_19"
   TextField "文本域_7" at 562,420 size 73x20; Text '设备正常'
   IOField "I/O 域_1" at 369,105 size 120x35; FormatPattern FFFFFFFF
      ProcessValue <- "故障代码x"
   IOField "I/O 域_2" at 623,255 size 120x35; FormatPattern FFFFFFFF
      ProcessValue <- "故障代码z"
   IOField "I/O 域_3" at 302,404 size 120x35; FormatPattern FFFFFFFF
      ProcessValue <- "故障代码y"
   TextField "文本域_8" at 703,356 size 73x20; Text '触发限位'
   Button "HmiScreenItemData_1" at 371,192 size 181x57; TextOff '伺服错误复位'; PictureOn "图形_13"; PictureOff "图形_38"
      on Release: ResetBit("HMI_MU_HMI伺服错误复位")
      on Press: SetBit("HMI_MU_HMI伺服错误复位")
   IOField "I/O 域_4" at 369,71 size 120x35; FormatPattern s9999.999; Unit MM
      ProcessValue <- "HengKongMC_hengkong_DATA_获取X轴当前坐标"
   IOField "I/O 域_5" at 623,221 size 120x35; FormatPattern s9999.999; Unit MM
      ProcessValue <- "HengKongMC_hengkong_DATA_获取Y轴当前坐标"
   IOField "I/O 域_6" at 302,369 size 120x35; FormatPattern s9999.999; Unit MM
      ProcessValue <- "HengKongMC_hengkong_DATA_获取Z轴当前坐标"
   TextField "文本域_9" at 24,67 size 19x29; Text 'X'
   TextField "文本域_10" at 24,125 size 19x29; Text 'Y'
   TextField "文本域_11" at 24,183 size 19x29; Text 'Z'

screen "补螺丝功能" 800x480, template "按钮_1"
   IOField "I/O 域_4" at 230,142 size 134x38; FormatPattern s999
      ProcessValue <- "HengKongMC_hengkong_报警异常号"
   IOField "I/O 域_6" at 230,230 size 134x38; FormatPattern s999
      ProcessValue <- "HengKongMC_hengkong_当前程序所在行号"
   Button "按钮_1" at 428,232 size 135x35; TextOff '写入'
      on Release: ResetBit("HengKongMC_hengkong_补螺丝功能_写入")
      on Press: SetBit("HengKongMC_hengkong_补螺丝功能_写入")
   Button "按钮_2" at 429,142 size 135x35; TextOff '读取'
      on Release: ResetBit("HengKongMC_hengkong_补螺丝功能_读取")
      on Press: SetBit("HengKongMC_hengkong_补螺丝功能_读取")
   Button "按钮_3" at 429,334 size 135x35; TextOff '从当前设定位置'
      on Release: SetTag("HengKongMC_hengkong_光标处运行标志", 1)
      Appearance <- "HengKongMC_hengkong_光标处运行标志"
   Button "按钮_4" at 229,334 size 135x35; TextOff '从第一行'
      on Release: SetTag("HengKongMC_hengkong_光标处运行标志", 0)
      Appearance <- "HengKongMC_hengkong_光标处运行标志"
   TextField "文本域_1" at 230,111 size 185x23; Text '当前锁螺丝错误行号'
   TextField "文本域_6" at 230,199 size 125x23; Text '设定错误行号'

screen "屏蔽管理_1" 800x480, template "按钮"
   Group "Group" at 359,67 size 422x401
   GraphicView "图形视图_2" at 159,305 size 50x50; Picture "图形_2"
   TextField "文本域_6" at 375,122 size 85x23; Text '光幕屏蔽'
   TextField "文本域_4" at 375,174 size 105x23; Text '安全门屏蔽'
   TextField "文本域_8" at 410,381 size 16x23; Text 'Text'
   SymbolicIOField "符号 I/O 域_1" at 595,113 size 157x32; TextOn '1'; TextOff '0'; TextList "屏蔽信号"
      ProcessValue <- "Blocking function_光幕屏蔽"
   SymbolicIOField "符号 I/O 域_2" at 595,165 size 157x32; TextOn '1'; TextOff '0'; TextList "屏蔽信号"
      ProcessValue <- "Blocking function_安全门屏蔽"
   SymbolicIOField "符号 I/O 域_8" at 185,69 size 160x35; TextOn '1'; TextOff '0'; TextList "屏蔽菜单"
      ProcessValue <- "屏蔽菜单"
      on Change: ActivateScreenByNumber("屏蔽菜单", 0)
   TextField "文本域_3" at 639,76 size 73x20; Text '操作按钮'
   TextField "文本域_2" at 421,76 size 73x20; Text '注释名称'

screen "报警历史" 800x480, template "按钮_1"
   AlarmView "报警视图_1" at 218,63 size 572x410; AlarmLog "报警历史"
   GraphicView "图形视图_2" at 153,244 size 50x50; Picture "图形_2"

screen "系统设置" 800x480, template "按钮_1"
   IOField "I/O 域_1" at 199,100 size 216x32; FormatPattern 9999999999999999999999999999999999999999
      ProcessValue <- "系统时间_WRDT"
   IOField "I/O 域_2" at 199,157 size 216x32; FormatPattern 9999999999999999999999999999999999999999
      ProcessValue <- "系统时间_RDDT"
   Button "按钮_1" at 420,100 size 96x32; TextOff '设置'
      on Press: SetBit("系统时间_SET")
      on Release: ResetBit("系统时间_SET")
   GraphicView "图形视图_7" at 159,374 size 50x50; Picture "图形_2"
   TextField "文本域_6" at 199,77 size 85x23; Text '设置时间'
   TextField "文本域_1" at 199,133 size 85x23; Text '系统时间'
   Button "HmiScreenItemData_5" at 639,406 size 143x47; TextOn '停止系统'; TextOff '关闭界面'; PictureOff "图形_21"; PictureOn "图形_21"
      on Release: StopRuntime(0)
*)